   IF #TankData.Active THEN
       CASE #TankData.TankState OF
           #TankState_Init:
               // This state is managed by the top level sequencer, no tank actions are required in this tank state.
               #TankData.XeOx_Complete := False;
               #TankData.Timer_Complete := False;
           #TankState_PreDwell:
               // This state is managed by the top level sequencer, no tank actions are required in this tank state.
               #TankData.XeOx_Complete := False;
               #TankData.Timer_Complete := False;
           #TankState_DeOx:
               CASE #State.DeOx OF
                   #State_DeOx_ClosePVV:
                       #PVVX_IN.PVVx_Actuate[#TankData.TankID] := True;
                       #PVVX_IN.PVVB_ValveDemands[#TankData.TankID] := False;
                       #PVVX_IN.PVVB_ValveDemands[#TankData.TankID] := False;
                   #State_DeOx_OpenGTT:
                       #GTT_IN.GTT_Actuate[#TankData.TankID] := True;
                       #GTT_IN.GTT_ValveDemands[#TankData.TankID] := True;
                       // Reset monitor timer in preparation for next stage
                       #MONITOR_TIMER(IN := False,
                                      PT := "1190_FIXED_CONSTANTS".DeOxAtLevel_Time,
                                      R := True);
                       #TankData.XeOx_Complete := False;
                   #State_DeOx_Monitor:
                       IF #MONITOR_TIMER.Q THEN
                           // Monitoring is complete, report this back to top level sequencer.
                           #TankData.XeOx_Complete := True;
                       ELSE
                           // Monitoring ongoing, check how to DO level compares to target,
                           // adjust the timer as appropriate (BWMS-100)
                           #TankData.XeOx_Complete := False;
                           IF #TankIPData.BWT_DO <= "1190_FIXED_CONSTANTS".DeOxTargetDOLevel THEN
                               // Tank DO level is equal or under target level, keep timer counting
                               #MONITOR_TIMER(IN := True,
                                              PT := "1190_FIXED_CONSTANTS".DeOxAtLevel_Time,
                                              R := False);
                           ELSE
                               // DO level has gone above target level. Reset the timer back to zero.
                               #MONITOR_TIMER(IN := False,
                                              PT := "1190_FIXED_CONSTANTS".DeOxAtLevel_Time,
                                              R := True);
                           END_IF;
                       END_IF;
                   #State_DeOx_CloseGTT:
                       #GTT_IN.GTT_Actuate[#TankData.TankID] := True;
                       #GTT_IN.GTT_ValveDemands[#TankData.TankID] := False;
                       // Reset the timer ready for Mid-Dwell phase
                       #DWELL_TIMER(IN := False,
                                    PT := "1190_FIXED_CONSTANTS".MidDwell_Time,
                                    R := True);
                       #TankData.Timer_Complete := false;
                   ELSE:
                       // another state in DeOx such as Start or Stop Supply to deck, no sub tank action is required as this is managed by the top level sequencer.
                       #TankData.XeOx_Complete := False;
                       #TankData.Timer_Complete := False;
               END_CASE;
           #TankState_MidDwell:
               // If this tank is in treatment group 1, update the middwell elapsed time so that the HMI
               // can be informed of the remaining time before the GCU needs to be activeated (BWMS-127,-128)
               IF (#State.TreatmentGroup = 1) THEN
                   "1191_SYSTEM_VARIABLES".MidDwell_ElapsedTime := #DWELL_TIMER.ET;
               END_IF;
               IF #DWELL_TIMER.Q THEN
                   #TankData.Timer_Complete := True;
               ELSE
                   #TankData.Timer_Complete := False;
                   // BWT DO level needs to remain under High DO Setpoint (BWMS-126)
                   IF #TankIPData.BWT_DO < "1094_ANALOGUE_SENSOR_SETPOINTS".TX427_428_DEOX.High THEN
                       #DWELL_TIMER(IN := True,
                                    PT := "1190_FIXED_CONSTANTS".MidDwell_Time,
                                    R := False);
                   ELSE
                       #DWELL_TIMER(IN := False,
                                    PT := "1190_FIXED_CONSTANTS".MidDwell_Time,
                                    R := True);
                   END_IF;
               END_IF;
           #TankState_ReOx:
               CASE #State.ReOx OF
                   #State_DwellAndReOx_OpenPVV:
                       #PVVX_IN.PVVx_Actuate[#TankData.TankID] := True;
                       #PVVX_IN.PVVB_ValveDemands[#TankData.TankID] := True;
                       #PVVX_IN.PVVB_ValveDemands[#TankData.TankID] := True;
                   #State_DwellAndReOx_OpenGTT:
                       #GTT_IN.GTT_Actuate[#TankData.TankID] := True;
                       #GTT_IN.GTT_ValveDemands[#TankData.TankID] := True;
                       // Reset monitor timer in preparation for next stage
                       #MONITOR_TIMER(IN := False,
                                      PT := "1190_FIXED_CONSTANTS".ReOxAtLevel_Time,
                                      R := True);
                       #ReOx_InitialTargetpHLevelAchieved := False;
                       #TankData.XeOx_Complete := False;
                   #State_DwellAndReOx_Monitor:
                       IF #MONITOR_TIMER.Q THEN
                           // Monitoring is complete, report this back to top level sequencer.
                           #TankData.XeOx_Complete := True;
                       ELSE
                           IF #ReOx_InitialTargetpHLevelAchieved THEN
                               // Monitoring ongoing, check how to pH level compares to low SP,
                               // adjust the timer as appropriate (BWMS-109)
                               #TankData.XeOx_Complete := False;
                               IF #TankIPData.BWT_PH > "1094_ANALOGUE_SENSOR_SETPOINTS".TX425_426.Low THEN
                                   // Tank pH level is greater than low SP, keep timer counting
                                   #MONITOR_TIMER(IN := True,
                                                  PT := "1190_FIXED_CONSTANTS".ReOxAtLevel_Time,
                                                  R := False);
                               ELSE
                                   // pH level has gone below or equal to low SP. Reset the timer back to zero.
                                   #MONITOR_TIMER(IN := False,
                                                  PT := "1190_FIXED_CONSTANTS".ReOxAtLevel_Time,
                                                  R := True);
                               END_IF;
                           ELSIF #TankIPData.BWT_PH >= "1190_FIXED_CONSTANTS".ReOxTargetpHLevel THEN
                               // Target level has been reached, timer started on next cycle, low SP then maintains timer reset.
                               #ReOx_InitialTargetpHLevelAchieved := true;
                           ELSE
                               // Target pH level has not been reached yet, keep timer in reset.
                               #MONITOR_TIMER(IN := False,
                                              PT := "1190_FIXED_CONSTANTS".ReOxAtLevel_Time,
                                              R := True);
                           END_IF;
                       END_IF;
                   #State_DwellAndReOx_CloseGTT:
                       #GTT_IN.GTT_Actuate[#TankData.TankID] := True;
                       #GTT_IN.GTT_ValveDemands[#TankData.TankID] := False;
                       // Reset dwell timer for next phase.
                       #TankData.Timer_Complete := False;
                       #DWELL_TIMER(IN := False,
                                    PT := "1190_FIXED_CONSTANTS".PostDwell_Time,
                                    R := True);
                   ELSE:
                       // another state in ReOx such as Start or Stop Supply to deck, no sub tank action is required as this is managed by the top level sequencer.
                       #TankData.XeOx_Complete := False;
                       #TankData.Timer_Complete := False;
               END_CASE;
           #TankState_PostDwell:
               // do timer functions wrt requirements
               IF #DWELL_TIMER.Q THEN
                   #TankData.Timer_Complete := True;
               ELSE
                   #TankData.Timer_Complete := False;
                   #DWELL_TIMER(IN := True,
                                PT := "1190_FIXED_CONSTANTS".PostDwell_Time,
                                R := False);
               END_IF;
           #TankState_Done:
               // Tank is complete, no further actions requried.
               #TankData.XeOx_Complete := False;
               #TankData.Timer_Complete := False;
       END_CASE;
   END_IF;
END_FUNCTION_BLOCK

// folder: 1000 - 1999 BWT System Control/1110 - 1129 Valve Control

FUNCTION_BLOCK "1110_DECK_MANAGE_START_SUPPLY"   // FB1110, SCL
{ S7_Optimized_Access := 'TRUE' }
VERSION : 0.1
   VAR RETAIN
      Stage : Int;
   END_VAR
   VAR
      DNC_500CV406 : "1604_DEMAND_AND_CHECK";
      DNC_600CV407 : "1604_DEMAND_AND_CHECK";
      DNC_600CV411 : "1604_DEMAND_AND_CHECK";
      DNC_600CV409 : "1604_DEMAND_AND_CHECK";
      TON_DELAY : TON_LTIME;
   END_VAR
   VAR RETAIN
      ShutdownDemand : Bool;
   END_VAR
BEGIN
   // Start the supply to the main deck. This is done in a specific order such that 
   // this operation is managed safely. If any stage fails the system will jump directly
   // to a shutdown state.

   CASE #Stage OF
       0:  // Reset all timers in Demand and check functions
           #DNC_500CV406.Reset := True;
           #DNC_500CV406.TRAVEL_TIME(IN := False,
                                     PT := LT#30s, // get real data from GCU code
                                     R := True);
           #DNC_600CV407.Reset := True;
           #DNC_600CV407.TRAVEL_TIME(IN := False,
                                     PT := "1096_ADJUSTABLE_CONSTANTS"."600CV407Open_Time",
                                     R := True);
           #DNC_600CV409.Reset := True;
           #DNC_600CV409.TRAVEL_TIME(IN := False,
                                     PT := "1096_ADJUSTABLE_CONSTANTS"."600CV409Close_time",
                                     R := True);
           #DNC_600CV411.Reset := True;
           #DNC_600CV411.TRAVEL_TIME(IN := False,
                                     PT := "1096_ADJUSTABLE_CONSTANTS"."600CV411Open_Time",
                                     R := True);
           #ShutdownDemand := False;
           #Stage += 1;
       1:  // Open Valve 500CV406 (NC)
           #DNC_500CV406.Reset := False;
           #DNC_500CV406(DemandIn := True,
                         NO_Type := False,
                         NC_Type := True,
                         ValveMoveTime := LT#30s,// get real data from GCU code
                         ValveOpenStatus := "10_DI_DATA".CV406_OPN,
                         ValveClsdStatus := "10_DI_DATA".CV406_CLSD,
                         DemandOut => "14_DQ_DATA".CV_406);
           IF #DNC_500CV406.DemandComplete AND NOT #DNC_500CV406.Alarm THEN
               #Stage += 1;
               #ShutdownDemand := false;
           ELSIF #DNC_500CV406.Alarm THEN
               #ShutdownDemand := true;
           END_IF;
           "1092_HMI_OP_FLAGS".DeckSupplyOk := False;
       2:  // Open Valve 600CV407 (NC)
           #DNC_600CV407.Reset := False;
           #DNC_600CV407(DemandIn := True,
                         NO_Type:=False,
                         NC_Type:=True,
                         ValveMoveTime:="1096_ADJUSTABLE_CONSTANTS"."600CV407Open_Time",
                         ValveOpenStatus := "10_DI_DATA".CV407_OPN,
                         ValveClsdStatus := "10_DI_DATA".CV407_CLSD,
                         DemandOut => "14_DQ_DATA".CV_407);
           IF #DNC_600CV407.DemandComplete AND NOT #DNC_600CV407.Alarm THEN
               #Stage += 1;
               #ShutdownDemand := false;
           ELSIF #DNC_600CV407.Alarm THEN
               #ShutdownDemand := true;
           END_IF;
           "1092_HMI_OP_FLAGS".DeckSupplyOk := False;
       3:  // Open Valve 600CV411 (NC)
           #DNC_600CV411.Reset := False;
           #DNC_600CV411(DemandIn := True,
                         NO_Type:=False,
                         NC_Type:=True,
                         ValveMoveTime:="1096_ADJUSTABLE_CONSTANTS"."600CV411Open_Time",
                         ValveOpenStatus := "10_DI_DATA".CV411_OPN,
                         ValveClsdStatus := "10_DI_DATA".CV411_CLSD,
                         DemandOut => "14_DQ_DATA".CV_411);
           IF #DNC_600CV411.DemandComplete AND NOT #DNC_600CV411.Alarm THEN
               #Stage += 1;
               #ShutdownDemand := false;
           ELSIF #DNC_600CV411.Alarm THEN
               #ShutdownDemand := true;
           END_IF;
           "1092_HMI_OP_FLAGS".DeckSupplyOk := False;
       4:  // Close 600CV409 (NO)
           #DNC_600CV409.Reset := False;
           #DNC_600CV409(DemandIn := True,
                         NO_Type:=True,
                         NC_Type:=False,
                         ValveMoveTime:="1096_ADJUSTABLE_CONSTANTS"."600CV409Close_time",
                         ValveOpenStatus := "10_DI_DATA".CV409_OPN,
                         ValveClsdStatus := "10_DI_DATA".CV409_CLSD,
                         DemandOut => "14_DQ_DATA".CV_409);
           IF #DNC_600CV409.DemandComplete AND NOT #DNC_600CV409.Alarm THEN
               #Stage += 1;
               #ShutdownDemand := false;
           ELSIF #DNC_600CV409.Alarm THEN
               #ShutdownDemand := true;
           END_IF;
           "1092_HMI_OP_FLAGS".DeckSupplyOk := False;
           #TON_DELAY(IN := false, // Reset the TON timer.
                      PT := T#15s);
       5:  // Wait for 15 seconds delay
           #TON_DELAY(IN := true,
                      PT := LT#15s);
           IF #TON_DELAY.Q THEN
               #Stage += 1;
               #TON_DELAY(IN := false, // Reset the TON timer for PIT415Delay_Time check
                          PT := T#15s);
           END_IF;
           "1092_HMI_OP_FLAGS".DeckSupplyOk := False;
           #ShutdownDemand := False;
       6:   // PIT415Delay_Time check of alarms.
           #TON_DELAY(IN := true,
                      PT := ("1096_ADJUSTABLE_CONSTANTS".PIT415Delay_Time - LT#15s));
           IF #TON_DELAY.Q AND NOT (#DNC_500CV406.Alarm OR #DNC_600CV407.Alarm OR #DNC_600CV409.Alarm OR #DNC_600CV411.Alarm) THEN
               // Supply is now ready, no alarms, end of process.
               "1092_HMI_OP_FLAGS".DeckSupplyOk := True;
               #ShutdownDemand := False;
           ELSIF (#DNC_500CV406.Alarm OR #DNC_600CV407.Alarm OR #DNC_600CV409.Alarm OR #DNC_600CV411.Alarm) THEN
               // Alarm raised, call shutdown
               #ShutdownDemand := True;
               "1092_HMI_OP_FLAGS".DeckSupplyOk := False;
           ELSE
               "1092_HMI_OP_FLAGS".DeckSupplyOk := False;
           END_IF;
       ELSE:
           // Unreachable branch - report error if reached.
           "1092_HMI_OP_FLAGS".DeckSupplyOk := False;
           #ShutdownDemand := True;
   END_CASE;
END_FUNCTION_BLOCK

FUNCTION_BLOCK "1111_DECK_MANAGE_STOP_SUPPLY"   // FB1111, SCL
{ S7_Optimized_Access := 'TRUE' }
VERSION : 0.1
   VAR RETAIN
      Stage : Int;
   END_VAR
   VAR
      DNC_500CV406 : "1604_DEMAND_AND_CHECK";
      DNC_600CV407 : "1604_DEMAND_AND_CHECK";
      DNC_600CV411 : "1604_DEMAND_AND_CHECK";
      DNC_600CV409 : "1604_DEMAND_AND_CHECK";
   END_VAR
   VAR RETAIN
      TON_DELAY : TON_TIME;
      ShutdownDemand : Bool;
      StopDeckSupplyDone : Bool;
   END_VAR
BEGIN
   // Stop the supply to the main deck. This is done in a specific order such that 
   // this operation is managed safely. If any stage fails the system will jump directly
   // to a shutdown state.

   CASE #Stage OF
       0:  // Reset all timers in Demand and check functions
           #DNC_500CV406.Reset := True;
           #DNC_500CV406.TRAVEL_TIME(IN := False,
                                     PT := LT#30s, // get real data from GCU code
                                     R := True);
           #DNC_600CV407.Reset := True;
           #DNC_600CV407.TRAVEL_TIME(IN := False,
                                     PT := "1096_ADJUSTABLE_CONSTANTS"."600CV407Close_Time",
                                     R := True);
           #DNC_600CV409.Reset := True;
           #DNC_600CV409.TRAVEL_TIME(IN := False,
                                     PT := "1096_ADJUSTABLE_CONSTANTS"."600CV409Open_Time",
                                     R := True);
           #DNC_600CV411.Reset := True;
           #DNC_600CV411.TRAVEL_TIME(IN := False,
                                     PT := "1096_ADJUSTABLE_CONSTANTS"."600CV411Close_time",
                                     R := True);
           #ShutdownDemand := False;
           "1092_HMI_OP_FLAGS".DeckSupplyOk := False;
           #StopDeckSupplyDone := False;
           #Stage += 1;
       1:  // Open Valve 600CV409 (NO)
           #DNC_600CV409.Reset := False;
           #DNC_600CV409(DemandIn := False,
                         NO_Type := True,
                         NC_Type := False,
                         ValveMoveTime := "1096_ADJUSTABLE_CONSTANTS"."600CV409Open_Time",
                         ValveClsdStatus := "10_DI_DATA".CV409_CLSD,
                         ValveOpenStatus := "10_DI_DATA".CV409_OPN,
                         DemandOut => "14_DQ_DATA".CV_409);
           IF #DNC_600CV409.DemandComplete AND NOT #DNC_600CV409.Alarm THEN
               #Stage += 1;
               #ShutdownDemand := false;
           ELSIF #DNC_600CV409.Alarm THEN
               #ShutdownDemand := true;
           END_IF;
           "1092_HMI_OP_FLAGS".DeckSupplyOk := False;
           #StopDeckSupplyDone := False;
       2:  // Close Valve 500CV406 (NC)
           #DNC_500CV406.Reset := False;
           #DNC_500CV406(DemandIn := False,
                         NO_Type := False,
                         NC_Type := True,
                         ValveMoveTime := T#30s, // get real data from GCU code
                         ValveClsdStatus := "10_DI_DATA".CV406_CLSD,
                         ValveOpenStatus := "10_DI_DATA".CV406_OPN,
                         DemandOut => "14_DQ_DATA".CV_406);
           IF #DNC_500CV406.DemandComplete AND NOT #DNC_500CV406.Alarm THEN
               #Stage += 1;
               #ShutdownDemand := false;
           ELSIF #DNC_500CV406.Alarm THEN
               #ShutdownDemand := true;
           END_IF;
           "1092_HMI_OP_FLAGS".DeckSupplyOk := False;
           #StopDeckSupplyDone := False;
       3: // Close Valve 600CV407 (NC)
           #DNC_600CV407.Reset := False;
           #DNC_600CV407(DemandIn := False,
                         NO_Type := False,
                         NC_Type := True,
                         ValveMoveTime := "1096_ADJUSTABLE_CONSTANTS"."600CV407Close_Time",
                         ValveClsdStatus := "10_DI_DATA".CV407_CLSD,
                         ValveOpenStatus := "10_DI_DATA".CV407_OPN,
                         DemandOut => "14_DQ_DATA".CV_407);
           IF #DNC_600CV407.DemandComplete AND NOT #DNC_600CV407.Alarm THEN
               #Stage += 1;
               #ShutdownDemand := false;
           ELSIF #DNC_600CV407.Alarm THEN
               #ShutdownDemand := true;
           END_IF;
           "1092_HMI_OP_FLAGS".DeckSupplyOk := False;
           #StopDeckSupplyDone := False;
       4: // Close Valve 600CV411 (NC)
           #DNC_600CV411.Reset := False;
           #DNC_600CV411(DemandIn := False,
                         NO_Type:=False,
                         NC_Type:=True,
                         ValveMoveTime:="1096_ADJUSTABLE_CONSTANTS"."600CV411Close_time",
                         ValveClsdStatus := "10_DI_DATA".CV411_CLSD,
                         ValveOpenStatus := "10_DI_DATA".CV411_OPN,
                         DemandOut => "14_DQ_DATA".CV_407);
           IF #DNC_600CV411.DemandComplete AND NOT #DNC_600CV411.Alarm THEN
               #Stage += 1;
               #ShutdownDemand := false;
           ELSIF #DNC_600CV411.Alarm THEN
               #ShutdownDemand := true;
           END_IF;
           "1092_HMI_OP_FLAGS".DeckSupplyOk := False;
           #StopDeckSupplyDone := False;
       5:  // Valves are now set.
           "1092_HMI_OP_FLAGS".DeckSupplyOk := False;
           #StopDeckSupplyDone := True;
       ELSE:
           // Unreachable branch - report error if reached.
           #StopDeckSupplyDone := False;
           #ShutdownDemand := True;
   END_CASE;
END_FUNCTION_BLOCK

FUNCTION_BLOCK "1115_GTT_MANAGE_VALVES"   // FB1115, LAD
{ S7_Optimized_Access := 'TRUE' }
VERSION : 0.1
// Manage the GTT (Gas To Tank/Inlet) valves based on the provided data.
// "Actuate" enables the actuation of the valves in question.
// "ValveDemands" signifies whether the valve should be actuating (Openning as NC valve) or releasing (Closing as NC valve).
// 
// This function puts out two sets of data:
// "DemandsCompleted" which indicates whether the demand is complete.
// "Alarms" indicated if an alarm has been triggered (e.g. a timeout in the Demand And Check.
// 
// The timeout for Demand and Check is automatically selected based on the demand and valve type.
   VAR_INPUT
      GTT_IN : "VALVE_GTT_IN";
   END_VAR
   VAR_IN_OUT
      GTT_OUT : "VALVE_GTT_OUT";
      GTT_Exclusivity : "GTT_EXCLUSIVITY";
   END_VAR
   VAR
      DNC_FPT_GTT : "1604_DEMAND_AND_CHECK";
      DNC_1P_GTT : "1604_DEMAND_AND_CHECK";
      DNC_1S_GTT : "1604_DEMAND_AND_CHECK";
      DNC_2P_GTT : "1604_DEMAND_AND_CHECK";
      DNC_2S_GTT : "1604_DEMAND_AND_CHECK";
      DNC_3P_GTT : "1604_DEMAND_AND_CHECK";
      DNC_3S_GTT : "1604_DEMAND_AND_CHECK";
      DNC_4P_GTT : "1604_DEMAND_AND_CHECK";
      DNC_4S_GTT : "1604_DEMAND_AND_CHECK";
      DNC_5P_GTT : "1604_DEMAND_AND_CHECK";
      DNC_5S_GTT : "1604_DEMAND_AND_CHECK";
      DNC_6P_GTT : "1604_DEMAND_AND_CHECK";
      DNC_6S_GTT : "1604_DEMAND_AND_CHECK";
      DNC_APT_GTT : "1604_DEMAND_AND_CHECK";
   END_VAR
   VAR_TEMP
      FPT_GTT_TimeSel : Time;
      "1P_GTT_TimeSel" : Time;
      "1S_GTT_TimeSel" : Time;
      "2P_GTT_TimeSel" : Time;
      "2S_GTT_TimeSel" : Time;
      "3P_GTT_TimeSel" : Time;
      "3S_GTT_TimeSel" : Time;
      "4P_GTT_TimeSel" : Time;
      "4S_GTT_TimeSel" : Time;
      "5P_GTT_TimeSel" : Time;
      "5S_GTT_TimeSel" : Time;
      "6P_GTT_TimeSel" : Time;
      "6S_GTT_TimeSel" : Time;
      APT_GTT_TimeSel : Time;
   END_VAR
   VAR CONSTANT
      TimerResetHold : LTime := LT#30s;
   END_VAR
   VAR_TEMP   // added for the SCL form of the ladder/FBD networks
      _w1 : Bool;
      _w2 : Bool;
      _w3 : Bool;
      _w4 : Bool;
      _w5 : Bool;
      _w6 : Bool;
      _w7 : Bool;
      _w8 : Bool;
      _w9 : Bool;
   END_VAR
BEGIN

REGION Network 1: Reset all timers if they are not in actuation mode.
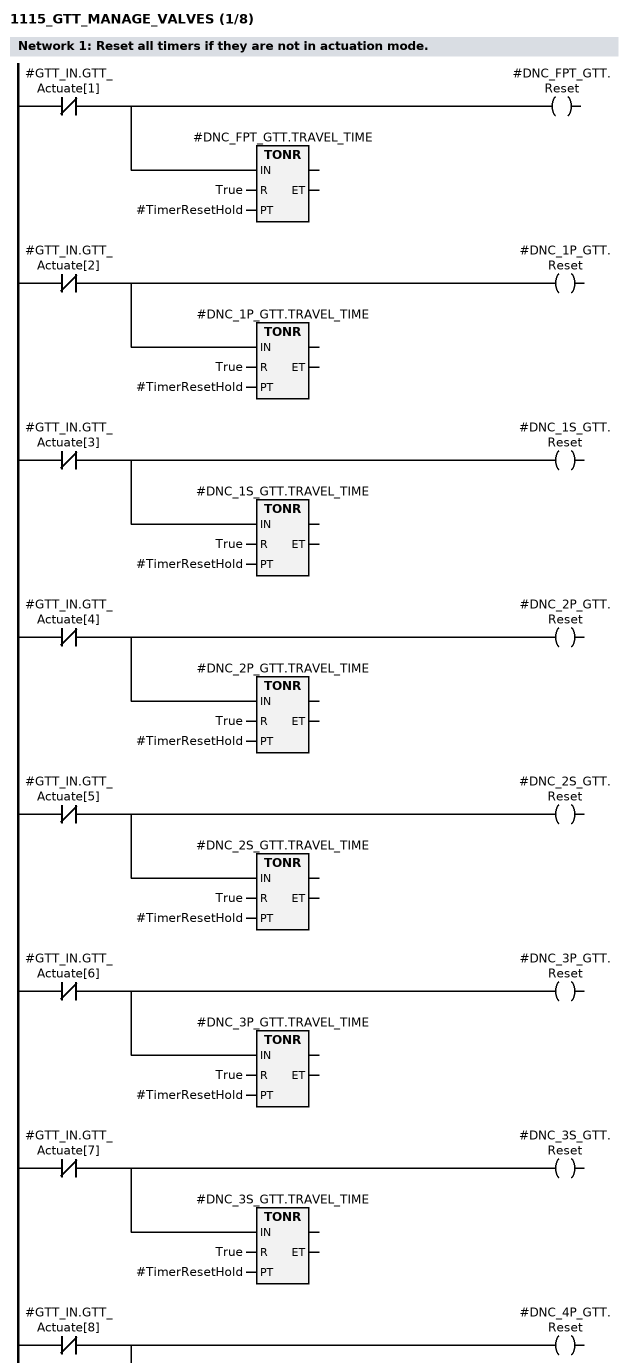
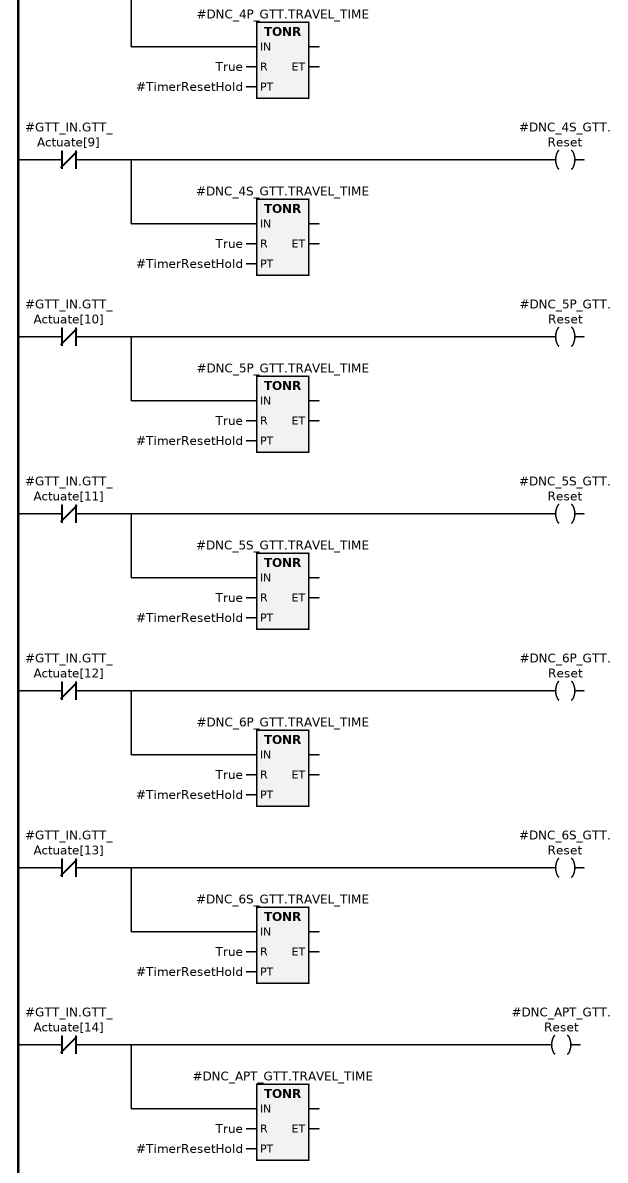
   #DNC_FPT_GTT.Reset := NOT #GTT_IN.GTT_Actuate[1];
   #DNC_FPT_GTT.TRAVEL_TIME.TONR(IN := NOT #GTT_IN.GTT_Actuate[1], R := True, PT := #TimerResetHold);
   #DNC_1P_GTT.Reset := NOT #GTT_IN.GTT_Actuate[2];
   #DNC_1P_GTT.TRAVEL_TIME.TONR(IN := NOT #GTT_IN.GTT_Actuate[2], R := True, PT := #TimerResetHold);
   #DNC_1S_GTT.Reset := NOT #GTT_IN.GTT_Actuate[3];
   #DNC_1S_GTT.TRAVEL_TIME.TONR(IN := NOT #GTT_IN.GTT_Actuate[3], R := True, PT := #TimerResetHold);
   #DNC_2P_GTT.Reset := NOT #GTT_IN.GTT_Actuate[4];
   #DNC_2P_GTT.TRAVEL_TIME.TONR(IN := NOT #GTT_IN.GTT_Actuate[4], R := True, PT := #TimerResetHold);
   #DNC_2S_GTT.Reset := NOT #GTT_IN.GTT_Actuate[5];
   #DNC_2S_GTT.TRAVEL_TIME.TONR(IN := NOT #GTT_IN.GTT_Actuate[5], R := True, PT := #TimerResetHold);
   #DNC_3P_GTT.Reset := NOT #GTT_IN.GTT_Actuate[6];
   #DNC_3P_GTT.TRAVEL_TIME.TONR(IN := NOT #GTT_IN.GTT_Actuate[6], R := True, PT := #TimerResetHold);
   #DNC_3S_GTT.Reset := NOT #GTT_IN.GTT_Actuate[7];
   #DNC_3S_GTT.TRAVEL_TIME.TONR(IN := NOT #GTT_IN.GTT_Actuate[7], R := True, PT := #TimerResetHold);
   #DNC_4P_GTT.Reset := NOT #GTT_IN.GTT_Actuate[8];
   #DNC_4P_GTT.TRAVEL_TIME.TONR(IN := NOT #GTT_IN.GTT_Actuate[8], R := True, PT := #TimerResetHold);
   #DNC_4S_GTT.Reset := NOT #GTT_IN.GTT_Actuate[9];
   #DNC_4S_GTT.TRAVEL_TIME.TONR(IN := NOT #GTT_IN.GTT_Actuate[9], R := True, PT := #TimerResetHold);
   #DNC_5P_GTT.Reset := NOT #GTT_IN.GTT_Actuate[10];
   #DNC_5P_GTT.TRAVEL_TIME.TONR(IN := NOT #GTT_IN.GTT_Actuate[10], R := True, PT := #TimerResetHold);
   #DNC_5S_GTT.Reset := NOT #GTT_IN.GTT_Actuate[11];
   #DNC_5S_GTT.TRAVEL_TIME.TONR(IN := NOT #GTT_IN.GTT_Actuate[11], R := True, PT := #TimerResetHold);
   #DNC_6P_GTT.Reset := NOT #GTT_IN.GTT_Actuate[12];
   #DNC_6P_GTT.TRAVEL_TIME.TONR(IN := NOT #GTT_IN.GTT_Actuate[12], R := True, PT := #TimerResetHold);
   #DNC_6S_GTT.Reset := NOT #GTT_IN.GTT_Actuate[13];
   #DNC_6S_GTT.TRAVEL_TIME.TONR(IN := NOT #GTT_IN.GTT_Actuate[13], R := True, PT := #TimerResetHold);
   #DNC_APT_GTT.Reset := NOT #GTT_IN.GTT_Actuate[14];
   #DNC_APT_GTT.TRAVEL_TIME.TONR(IN := NOT #GTT_IN.GTT_Actuate[14], R := True, PT := #TimerResetHold);
END_REGION

REGION Network 2: RIO01 FPT, 1P, 1S GTT control
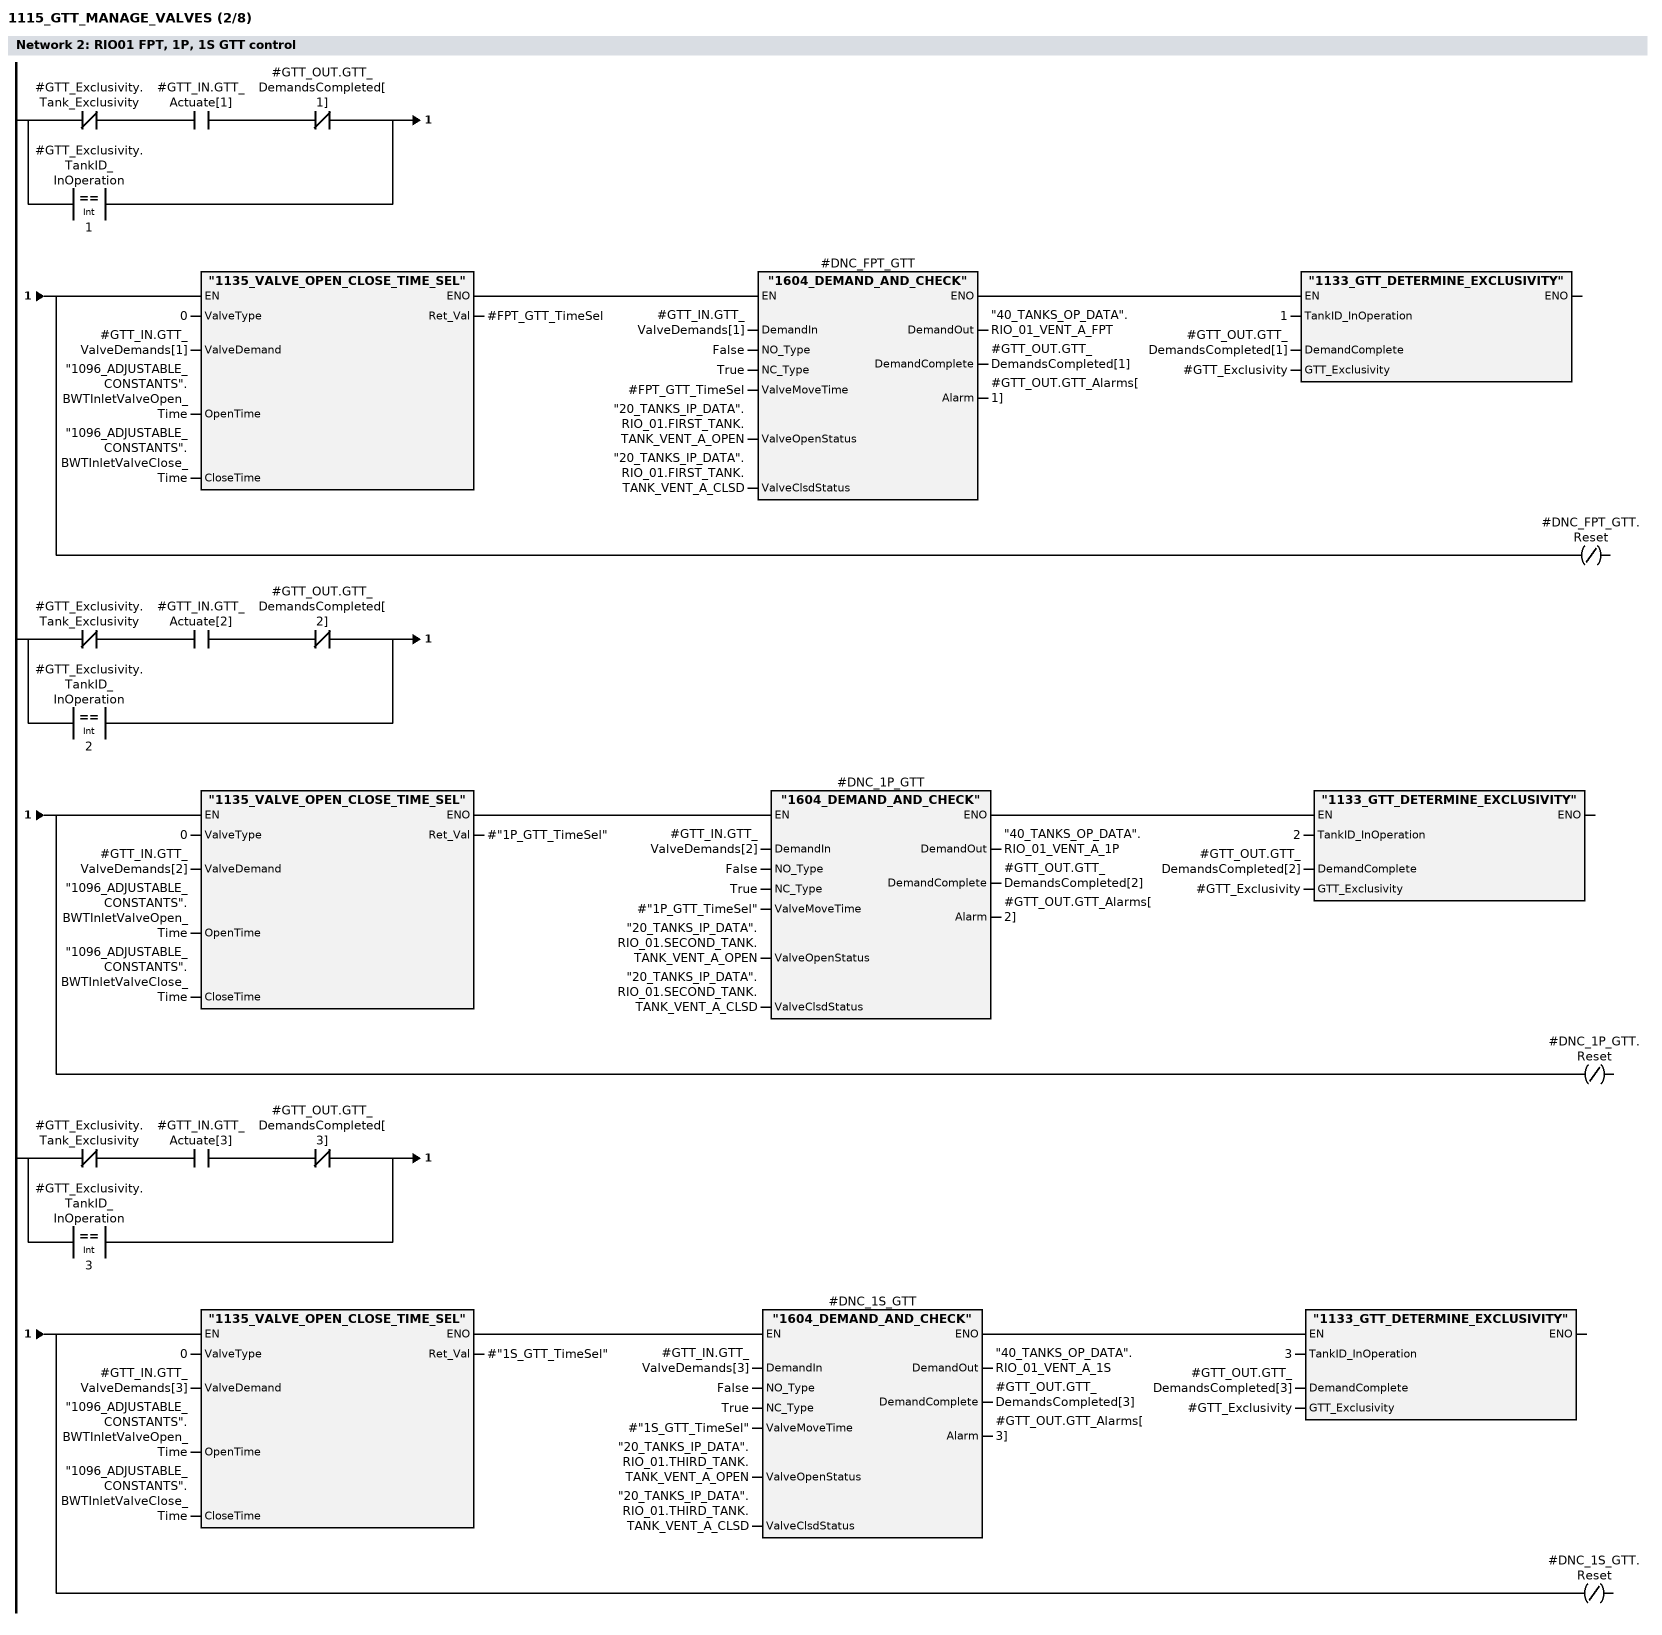
   RUNG wire#powerrail
      I_Contact( #GTT_Exclusivity.Tank_Exclusivity )
      Contact( #GTT_IN.GTT_Actuate[1] )
      I_Contact( #GTT_OUT.GTT_DemandsCompleted[1] )
      wire#w1
      "1135_VALVE_OPEN_CLOSE_TIME_SEL"(ValveType := 0, ValveDemand := #GTT_IN.GTT_ValveDemands[1], OpenTime := "1096_ADJUSTABLE_CONSTANTS".BWTInletValveOpen_Time, CloseTime := "1096_ADJUSTABLE_CONSTANTS".BWTInletValveClose_Time, Ret_Val => #FPT_GTT_TimeSel)
      #DNC_FPT_GTT(DemandIn := #GTT_IN.GTT_ValveDemands[1], NO_Type := False, NC_Type := True, ValveMoveTime := #FPT_GTT_TimeSel, ValveOpenStatus := "20_TANKS_IP_DATA".RIO_01.FIRST_TANK.TANK_VENT_A_OPEN, ValveClsdStatus := "20_TANKS_IP_DATA".RIO_01.FIRST_TANK.TANK_VENT_A_CLSD, DemandOut => "40_TANKS_OP_DATA".RIO_01_VENT_A_FPT, DemandComplete => #GTT_OUT.GTT_DemandsCompleted[1], Alarm => #GTT_OUT.GTT_Alarms[1])
      "1133_GTT_DETERMINE_EXCLUSIVITY"(TankID_InOperation := 1, DemandComplete := #GTT_OUT.GTT_DemandsCompleted[1], GTT_Exclusivity := #GTT_Exclusivity)
   END_RUNG
   RUNG wire#powerrail
      { S7_Templates := "SrcType := Int" } EQ_Contact(in1 := #GTT_Exclusivity.TankID_InOperation, in2 := 1)
   END_RUNG wire#w1
   RUNG wire#w1
      I_Coil( #DNC_FPT_GTT.Reset )
   END_RUNG
   RUNG wire#powerrail
      I_Contact( #GTT_Exclusivity.Tank_Exclusivity )
      Contact( #GTT_IN.GTT_Actuate[2] )
      I_Contact( #GTT_OUT.GTT_DemandsCompleted[2] )
      wire#w2
      "1135_VALVE_OPEN_CLOSE_TIME_SEL"(ValveType := 0, ValveDemand := #GTT_IN.GTT_ValveDemands[2], OpenTime := "1096_ADJUSTABLE_CONSTANTS".BWTInletValveOpen_Time, CloseTime := "1096_ADJUSTABLE_CONSTANTS".BWTInletValveClose_Time, Ret_Val => #"1P_GTT_TimeSel")
      #DNC_1P_GTT(DemandIn := #GTT_IN.GTT_ValveDemands[2], NO_Type := False, NC_Type := True, ValveMoveTime := #"1P_GTT_TimeSel", ValveOpenStatus := "20_TANKS_IP_DATA".RIO_01.SECOND_TANK.TANK_VENT_A_OPEN, ValveClsdStatus := "20_TANKS_IP_DATA".RIO_01.SECOND_TANK.TANK_VENT_A_CLSD, DemandOut => "40_TANKS_OP_DATA".RIO_01_VENT_A_1P, DemandComplete => #GTT_OUT.GTT_DemandsCompleted[2], Alarm => #GTT_OUT.GTT_Alarms[2])
      "1133_GTT_DETERMINE_EXCLUSIVITY"(TankID_InOperation := 2, DemandComplete := #GTT_OUT.GTT_DemandsCompleted[2], GTT_Exclusivity := #GTT_Exclusivity)
   END_RUNG
   RUNG wire#powerrail
      { S7_Templates := "SrcType := Int" } EQ_Contact(in1 := #GTT_Exclusivity.TankID_InOperation, in2 := 2)
   END_RUNG wire#w2
   RUNG wire#w2
      I_Coil( #DNC_1P_GTT.Reset )
   END_RUNG
   RUNG wire#powerrail
      I_Contact( #GTT_Exclusivity.Tank_Exclusivity )
      Contact( #GTT_IN.GTT_Actuate[3] )
      I_Contact( #GTT_OUT.GTT_DemandsCompleted[3] )
      wire#w3
      "1135_VALVE_OPEN_CLOSE_TIME_SEL"(ValveType := 0, ValveDemand := #GTT_IN.GTT_ValveDemands[3], OpenTime := "1096_ADJUSTABLE_CONSTANTS".BWTInletValveOpen_Time, CloseTime := "1096_ADJUSTABLE_CONSTANTS".BWTInletValveClose_Time, Ret_Val => #"1S_GTT_TimeSel")
      #DNC_1S_GTT(DemandIn := #GTT_IN.GTT_ValveDemands[3], NO_Type := False, NC_Type := True, ValveMoveTime := #"1S_GTT_TimeSel", ValveOpenStatus := "20_TANKS_IP_DATA".RIO_01.THIRD_TANK.TANK_VENT_A_OPEN, ValveClsdStatus := "20_TANKS_IP_DATA".RIO_01.THIRD_TANK.TANK_VENT_A_CLSD, DemandOut => "40_TANKS_OP_DATA".RIO_01_VENT_A_1S, DemandComplete => #GTT_OUT.GTT_DemandsCompleted[3], Alarm => #GTT_OUT.GTT_Alarms[3])
      "1133_GTT_DETERMINE_EXCLUSIVITY"(TankID_InOperation := 3, DemandComplete := #GTT_OUT.GTT_DemandsCompleted[3], GTT_Exclusivity := #GTT_Exclusivity)
   END_RUNG
   RUNG wire#powerrail
      { S7_Templates := "SrcType := Int" } EQ_Contact(in1 := #GTT_Exclusivity.TankID_InOperation, in2 := 3)
   END_RUNG wire#w3
   RUNG wire#w3
      I_Coil( #DNC_1S_GTT.Reset )
   END_RUNG
   // the same network as SCL:
   #_w1 := (NOT #GTT_Exclusivity.Tank_Exclusivity AND #GTT_IN.GTT_Actuate[1] AND NOT #GTT_OUT.GTT_DemandsCompleted[1]) OR (#GTT_Exclusivity.TankID_InOperation = 1);
   #FPT_GTT_TimeSel := "1135_VALVE_OPEN_CLOSE_TIME_SEL"(EN := #_w1,
                           ValveType := 0,